   // NTTS[55] := 57;
   // NTTS[56] := 58;
   // NTTS[57] := 59;
   // NTTS[58] := 60;
   // NTTS[59] := 61;
   // NTTS[60] := 62;
   // NTTS[61] := 63;
   // NTTS[62] := 64;
   // NTTS[63] := 66;
   // SW_SQTS[2] := 1;
   // SW_SQTS[8] := 2;
   // SW_SQTS[9] := 2;
   // SW_SQTS[10] := 3;
   // SW_SQTS[11] := 3;
   // SW_SQTS[12] := 3;
   // SW_SQTS[13] := 3;
   // SW_SQTS[14] := 4;
   // SW_SQTS[15] := 4;
   // SW_SQTS[16] := 4;
   // SW_SQTS[17] := 4;
   // SW_SQTS[18] := 4;
   // SW_SQTS[19] := 4;
   // SW_SQTS[20] := 5;
   // SW_SQTS[21] := 5;
   // SW_SQTS[22] := 5;
   // SW_SQTS[23] := 2;
   // SW_SQTS[24] := 6;
   // SW_SQTS[25] := 6;
   // SW_SQTS[26] := 6;
   // SW_SQTS[27] := 6;
   // SW_SQTS[28] := 6;
   // SW_SQTS[29] := 6;
   // SW_SQTS[30] := 6;
   // SW_SQTS[31] := 6;
   // SWITCH[3] := 240;
   // SW_SQTS[36] := 7;
   // SW_SQTS[37] := 7;
   // SW_SQTS[38] := 7;
   // SW_SQTS[39] := 7;
   // SW_SQTS[40] := 7;
   // SW_SQTS[41] := 7;
   // SW_SQTS[42] := 7;
   // SW_SQTS[43] := 7;
   // SW_SQTS[44] := 7;
   // SW_SQTS[45] := 8;
   // SW_SQTS[46] := 8;
   // SW_SQTS[47] := 8;
   // SW_SQTS[48] := 8;
   // SW_SQTS[49] := 8;
   // SW_SQTS[50] := 8;
   // SW_SQTS[51] := 8;
   // SW_SQTS[52] := 8;
   // SW_SQTS[53] := 8;
   // SW_SQTS[54] := 8;
   // SW_SQTS[55] := 8;
   // SW_SQTS[56] := 8;
   // SW_SQTS[57] := 8;
   // SW_SQTS[58] := 8;
   // SW_SQTS[59] := 9;
   // SW_SQTS[60] := 9;
   // SW_SQTS[61] := 9;
   // SW_SQTS[62] := 9;
   // SW_SQTS[63] := 10;
   // SWITCH[0] := 252;
   // SWITCH[8] := 255;
   // SWITCH[4] := 167;
   // SWITCH[5] := 191;
   // SWITCH[6] := 252;
   // SWITCH[7] := 225;
   // SWITCH[2] := 255;
   // NSTT[48] := 47;
   // PTTS[27] := 34;
   // NSTT[38] := 37;
   // PTTS[30] := 31;
   // NTTS[1] := 3;
   // SWITCH[14] := 255;
   // ATAB[20] := 20;
   // PSTT[11] := 7;
   // NTTS[2] := 4;
   // PTTS[4] := 26;
   // PTTS[1] := 2;
   // NTTS[4] := 8;
   // SW_SQTS[1] := 1;
   // NSTT[26] := 4;
   // LSTT[48] := 255;
   // LSTT[63] := 255;
   // NSTT[63] := 62;
   // LSTT[61] := 255;
   // NSTT[61] := 60;
   // LSTT[64] := 1;
   // NSTT[64] := 1;
   // "Aux Reactor"."TIMER".MIX.PT := T#5M;
   // "Aux Reactor"."TIMER"."PRE-MIX".PT := T#5M;
   // SINI[6] := 255;
   // "Aux Reactor"."TIMER".TUBE.PT := T#5M;
   // "Aux Reactor"."TIMER".WASH.PT := T#5M;
   // SINI[5] := 255;
   // "Aux Reactor"."TIMER".REACTOR.PT := T#21.5H;
   // "Aux Reactor"."TIMER".PH_DELAY.PT := T#1M;
   // PTTS[29] := 30;
   // LSTT[37] := 255;
   // LSTT[25] := 24;
   // ATAB[19] := 19;
   // PSTT[15] := 11;
   // NSTT[37] := 36;
   // NSTT[25] := 24;
   // PTTS[28] := 28;
   // SW_SQTS[7] := 2;
   // SW_SQTS[6] := 2;
   // SW_SQTS[5] := 2;
   // SW_SQTS[4] := 2;
   // SWITCH[11] := 255;
   // SWITCH[13] := 239;
   // SWITCH[12] := 254;
   // PSTT[34] := 32;
   // PSTT[55] := 53;
   // PSTT[54] := 52;
   // LSTT[26] := 255;
   // SWITCH[10] := 239;
   // SWITCH[9] := 254;
   // SWITCH[1] := 231;
   // PTTS[2] := 3;
   // NSTT[49] := 48;
   // PSTT[53] := 51;
   // ATAB[0] := 1;
   // LSTT[49] := 255;
   // SINI[4] := 255;
   // SINI[2] := 255;
   // SW_SQTS[33] := 6;
   // SW_SQTS[32] := 6;
   // SINI[7] := 255;
   // SINI[8] := 255;
   // SINI[9] := 255;
   // LSTT[34] := 255;
   // LSTT[43] := 255;
   // PSTT[39] := 37;
   // NSTT[43] := 43;
   // LSTT[28] := 255;
   // LSTT[33] := 255;
   // ATAJ[66] := 66;
   // ATAB[66] := 66;
   // PSTT[66] := 63;
   // NSTT[33] := 26;
   // ASSJ[64] := 64;
   // ASSB[64] := 64;
   // PTTS[64] := 66;
   // NTTS[64] := 67;
   // SW_SQTS[64] := 10;
   // ATAJ[67] := 67;
   // ATAB[67] := 67;
   // PSTT[67] := 64;
   // NSTT[34] := 27;
   // LSTT[67] := 255;
   // ATAJ[68] := 68;
   // ATAB[68] := 68;
   // PSTT[68] := 65;
   // NSTT[67] := 65;
   // ASSJ[65] := 65;
   // ASSB[65] := 65;
   // PTTS[65] := 67;
   // NTTS[65] := 68;
   // SW_SQTS[65] := 10;
BEGIN
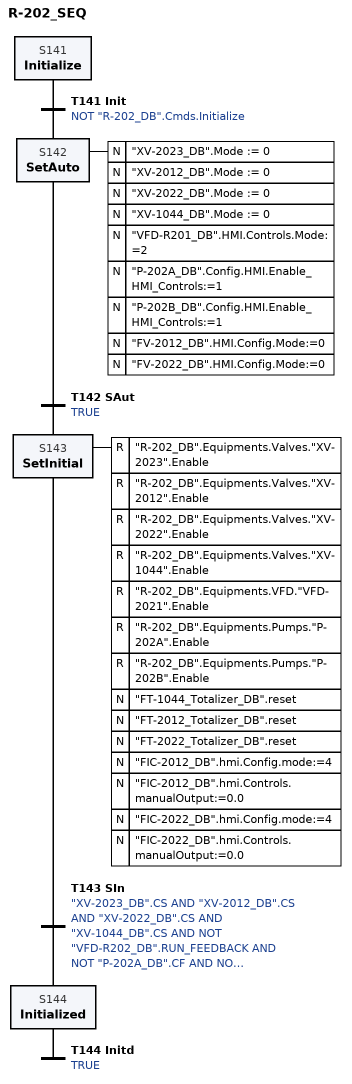
   // permanent pre-instructions
   NETWORK 1
      "R-202_Signals_FROM_T-101"();
      "R-202_Signals_FROM_T-102"();
      "R-202_Signals_FROM_T-103"();
      "R-202_Signals_FROM_T-104"();
      "R-202_SEQ_FC"();
      "R-202_Transitions_FC"();

   // sequencer 1
   STEP Initialize:   // S141, max time T#10S, warning time T#7S
   END_STEP
   TRANSITION Init FROM Initialize TO SetAuto   // T141
      := NOT "R-202_DB".Cmds.Initialize;
   END_TRANSITION
   STEP SetAuto:   // S142, max time T#10S, warning time T#7S
              N    "XV-2023_DB".Mode := 0
              N    "XV-2012_DB".Mode := 0
              N    "XV-2022_DB".Mode := 0
              N    "XV-1044_DB".Mode := 0
              N    "VFD-R201_DB".HMI.Controls.Mode:=2
              N    "P-202A_DB".Config.HMI.Enable_HMI_Controls:=1
              N    "P-202B_DB".Config.HMI.Enable_HMI_Controls:=1
              N    "FV-2012_DB".HMI.Config.Mode:=0
              N    "FV-2022_DB".HMI.Config.Mode:=0
   END_STEP
   TRANSITION SAut FROM SetAuto TO SetInitial   // T142
      := TRUE;
   END_TRANSITION
   STEP SetInitial:   // S143, max time T#10S, warning time T#7S
              R    "R-202_DB".Equipments.Valves."XV-2023".Enable
              R    "R-202_DB".Equipments.Valves."XV-2012".Enable
              R    "R-202_DB".Equipments.Valves."XV-2022".Enable
              R    "R-202_DB".Equipments.Valves."XV-1044".Enable
              R    "R-202_DB".Equipments.VFD."VFD-2021".Enable
              R    "R-202_DB".Equipments.Pumps."P-202A".Enable
              R    "R-202_DB".Equipments.Pumps."P-202B".Enable
              N    "FT-1044_Totalizer_DB".reset
              N    "FT-2012_Totalizer_DB".reset
              N    "FT-2022_Totalizer_DB".reset
              N    "FIC-2012_DB".hmi.Config.mode:=4
              N    "FIC-2012_DB".hmi.Controls.manualOutput:=0.0
              N    "FIC-2022_DB".hmi.Config.mode:=4
              N    "FIC-2022_DB".hmi.Controls.manualOutput:=0.0
   END_STEP
   TRANSITION SIn FROM SetInitial TO Initialized   // T143
      := "XV-2023_DB".CS AND "XV-2012_DB".CS AND "XV-2022_DB".CS AND "XV-1044_DB".CS AND NOT "VFD-R202_DB".RUN_FEEDBACK AND NOT "P-202A_DB".CF AND NOT "P-202B_DB".CF AND ("FV-2011_DB".CMD <= 0) AND ("FV-2021_DB".CMD <= 0) AND ("FT-1044_Totalizer_DB".Total = 0.0) AND ("FT-2012_Totalizer_DB".Total = 0.0) AND ("FT-2022_Totalizer_DB".Total = 0.0);
   END_TRANSITION
   STEP Initialized:   // S144, max time T#10S, warning time T#7S
      // Done Initialization
   END_STEP
   TRANSITION Initd FROM Initialized TO ?   // T144
      := TRUE;
   END_TRANSITION

   // permanent post-instructions
   NETWORK 1
      "R-202_FC_Outputs"();
END_FUNCTION_BLOCK

FUNCTION "R-202_FC_Outputs" : Void   // FC43, SCL
{ S7_Optimized_Access := 'TRUE' }
VERSION : 0.1
   VAR_TEMP
      Pump_A : Struct
         Cond_01 : Bool;   // Condition 01
         Cond_02 : Bool;
         Cond_03 : Bool;   // Condition 03
      END_STRUCT;
      Pump_B : Struct
         Cond_01 : Bool;   // Condition 01
         Cond_02 : Bool;   // Condition 02
         Cond_03 : Bool;   // Condition 03
      END_STRUCT;
      Motor : Struct
         Cond_01 : Bool;   // Condition 01
         Cond_02 : Bool;   // Condition 02
         Cond_03 : Bool;   // Condition 03
      END_STRUCT;
      XV : Struct
         "2023" : Bool;
         "2012" : Bool;
         "2022" : Bool;
         "1044" : Bool;
      END_STRUCT;
      "FV-2012" : Struct
         On : Bool;
         Cond_1 : Bool;
      END_STRUCT;
      "FV-2022" : Struct
         On : Bool;
         Cond_1 : Bool;
      END_STRUCT;
   END_VAR
BEGIN
   //****** Equipmens Activation*******
   //
   //**************************************************************
   //
   //IF "AlwaysFALSE" THEN
       //***********************************************Reactor Outlet Valve**********************************************************************
       IF "XV-2023_DB".Mode = 0 THEN
           "R-202_DB".Equipments.Valves."XV-2023".CmdOn := "R-202_DB".Equipments.Valves."XV-2023".Enable AND NOT "R-202_DB".Cmds.Hold;
           //Delay Off To avoid Overpressure the Lines
           #XV."2023" := "R-202_DB".Equipments.Valves."XV-2023".CmdOn;
           "R-202_Aux_DB".Timer."XV-2023".TOF(IN := #XV."2023",
                                              PT := "R-202_Aux_DB".Constants.CmdDelay);
           //Command to the Valve
           IF "R-202_Aux_DB".Timer."XV-2023".Q THEN
               "XV-2023_DB".CMD := 2;
           ELSE
               "XV-2023_DB".CMD := 1;
           END_IF;
           "R-202_DB".Equipments.Valves."XV-2023".TurningOff := NOT "R-202_DB".Equipments.Valves."XV-2023".CmdOn AND "R-202_Aux_DB".Timer."XV-2023".Q;
       END_IF;
       //***********************************************From T-101 Inlet Route********************************************************************
       IF "XV-2012_DB".Mode = 0 THEN
           "R-202_DB".Equipments.Valves."XV-2012".CmdOn := "R-202_DB".Equipments.Valves."XV-2012".Enable AND NOT "R-202_DB".Cmds.Hold;
           //Delay Off To avoid Overpressure the Lines
           #XV."2012" := "R-202_DB".Equipments.Valves."XV-2012".CmdOn;
           "R-202_Aux_DB".Timer."XV-2012".TOF(IN := #XV."2012",
                                              PT := "R-202_Aux_DB".Constants.CmdDelay);
           //Command to the Valve
           IF "R-202_Aux_DB".Timer."XV-2012".Q THEN
               "XV-2012_DB".CMD := 2;
           ELSE
               "XV-2012_DB".CMD := 1;
           END_IF;
           "R-202_DB".Equipments.Valves."XV-2012".TurningOff := NOT "R-202_DB".Equipments.Valves."XV-2012".CmdOn AND "R-202_Aux_DB".Timer."XV-2012".Q;
       END_IF;
       //***********************************************From T-102 Inlet Route********************************************************************
       IF "XV-2022_DB".Mode = 0 THEN
           "R-202_DB".Equipments.Valves."XV-2022".CmdOn := "R-202_DB".Equipments.Valves."XV-2022".Enable AND NOT "R-202_DB".Cmds.Hold;
           //Delay Off To avoid Overpressure the Lines
           #XV."2022" := "R-202_DB".Equipments.Valves."XV-2022".CmdOn;
           "R-202_Aux_DB".Timer."XV-2022".TOF(IN := #XV."2022",
                                              PT := "R-202_Aux_DB".Constants.CmdDelay);
           //Command to the Valve
           IF "R-202_Aux_DB".Timer."XV-2022".Q THEN
               "XV-2022_DB".CMD := 2;
           ELSE
               "XV-2022_DB".CMD := 1;
           END_IF;
           "R-202_DB".Equipments.Valves."XV-2022".TurningOff := NOT "R-202_DB".Equipments.Valves."XV-2022".CmdOn AND "R-202_Aux_DB".Timer."XV-2022".Q;
       END_IF;
       //***********************************************From T-104 Inlet Route (Water)********************************************************************
       IF "XV-1044_DB".Mode = 0 THEN
           "R-202_DB".Equipments.Valves."XV-1044".CmdOn := "R-202_DB".Equipments.Valves."XV-1044".Enable AND NOT "R-202_DB".Cmds.Hold;
           //Delay Off To avoid Overpressure the Lines
           #XV."1044" := "R-202_DB".Equipments.Valves."XV-1044".CmdOn;
           "R-202_Aux_DB".Timer."XV-1044".TOF(IN := #XV."1044",
                                              PT := "R-202_Aux_DB".Constants.CmdDelay);
           //Command to the Valve
           IF "R-202_Aux_DB".Timer."XV-1044".Q THEN
               "XV-1044_DB".CMD := 2;
           ELSE
               "XV-1044_DB".CMD := 1;
           END_IF;
           "R-202_DB".Equipments.Valves."XV-1044".TurningOff := NOT "R-202_DB".Equipments.Valves."XV-1044".CmdOn AND "R-202_Aux_DB".Timer."XV-2022".Q;
       END_IF;
       //***********************************************FIC-2012 Controller (From T-101)********************************************************************
       IF "FV-2012_DB".HMI.Config.Mode = 0 THEN
           #"FV-2012".Cond_1 := "R-202_DB".Equipments.Valves."FV-2012".Enable AND "XV-2012_DB".OS;
           "R-202_DB".Equipments.Valves."FV-2012".CmdOn := #"FV-2012".Cond_1 AND NOT "R-202_DB".Cmds.Hold AND NOT "R-202_DB".Status.Aborting;
           //Delay Off To avoid Overpressure the Lines
           #"FV-2012".On := "R-202_DB".Equipments.Valves."FV-2012".CmdOn;
           "R-202_Aux_DB".Timer."FV-2012".TOF(IN := #"FV-2012".On,
                                              PT := "R-202_Aux_DB".Constants.CmdDelay);
           IF "R-202_Aux_DB".Timer."FV-2012".Q THEN
               "FIC-2012_DB".enableManualMode := False;
               "FIC-2012_DB".enableRemoteSetpoint := False;
               "FIC-2012_DB".hmi.Controls.manualEnable := False;
               "FIC-2012_DB".hmi.Config.mode := 3;
           END_IF;     // ELSE
              // "FIC-2012_DB".enableManualMode := True;
              // "FIC-2012_DB".hmi.Controls.manualEnable := True;
              // "FIC-2012_DB".hmi.Config.mode := 4;
              // "FIC-2012_DB".hmi.Controls.manualOutput := 0;
         //  END_IF;
           "R-202_DB".Equipments.Valves."FV-2012".TurningOff := NOT "R-202_DB".Equipments.Valves."FV-2012".CmdOn AND "R-202_Aux_DB".Timer."FV-2012".Q;
       END_IF;
       //***********************************************FIC-2022 Controller (From T-102)********************************************************************
       IF "FV-2022_DB".HMI.Config.Mode = 0 THEN
           #"FV-2022".Cond_1 := "R-202_DB".Equipments.Valves."FV-2022".Enable AND "XV-2022_DB".OS;
           "R-202_DB".Equipments.Valves."FV-2022".CmdOn := #"FV-2022".Cond_1 AND NOT "R-202_DB".Cmds.Hold AND NOT "R-202_DB".Status.Aborting;
           //Delay Off To avoid Overpressure the Lines
           #"FV-2022".On := "R-202_DB".Equipments.Valves."FV-2022".CmdOn;
           "R-202_Aux_DB".Timer."FV-2022".TOF(IN := #"FV-2022".On,
                                              PT := "R-202_Aux_DB".Constants.CmdDelay);
           IF "R-202_Aux_DB".Timer."FV-2022".Q THEN

               IF "R-202_SEQ_DB".pH_Ctrl1.X OR "R-202_SEQ_DB".pH_Ctrl2.X OR "R-202_SEQ_DB".FillDone_T102.X THEN
                   //FIC-2022 Secondary Controller
                   "FIC-2022_DB".enableManualMode := False;
                   "FIC-2022_DB".hmi.Controls.manualEnable := False;
                   "FIC-2022_DB".enableRemoteSetpoint := true;
                   "FIC-2022_DB".hmi.Config.mode := 6;

                   //PHIC-R-202 pH Primary Controller
                   "PHIC-R-202_DB".enableRemoteSetpoint := False;
                   "PHIC-R-202_DB".enableManualMode := False;
                   "PHIC-R-202_DB".hmi.Controls.manualEnable := False;
                   "PHIC-R-202_DB".hmi.Config.mode := 3;
               ELSIF "R-202_SEQ_DB".Y.X THEN
                   //FIC-2022 Secondary Controller
                   "FIC-2022_DB".enableManualMode := False;
                   "FIC-2022_DB".hmi.Controls.manualEnable := False;
                   "FIC-2022_DB".enableRemoteSetpoint := false;
                   "FIC-2022_DB".hmi.Config.mode := 3;

                   //PHIC-R-202 pH Primary Controller
                   "PHIC-R-202_DB".enableRemoteSetpoint := False;
                   "PHIC-R-202_DB".enableManualMode := False;
                   "PHIC-R-202_DB".hmi.Controls.manualEnable := False;
                   "PHIC-R-202_DB".hmi.Config.mode := 3;

               END_IF;



           END_IF;     // ELSE
               //FIC-2022 Secondary Controller
             //  "FIC-2022_DB".enableManualMode := True;
             //  "FIC-2022_DB".hmi.Controls.manualEnable := True;
             //  "FIC-2022_DB".enableRemoteSetpoint := False;
             //  "FIC-2022_DB".hmi.Config.mode := 4;
             //  "FIC-2022_DB".hmi.Controls.manualOutput := 0;

               //PHIC-R-202 pH Primary  Controller
             //  "PHIC-R-202_DB".enableManualMode := True;
             //  "PHIC-R-202_DB".hmi.Controls.manualEnable := True;
             //  "PHIC-R-202_DB".enableRemoteSetpoint := False;
             //  "PHIC-R-202_DB".hmi.Config.mode := 4;
            //   "PHIC-R-202_DB".hmi.Controls.manualOutput := 0;
         //  END_IF;
           "R-202_DB".Equipments.Valves."FV-2022".TurningOff := NOT "R-202_DB".Equipments.Valves."FV-2022".CmdOn AND "R-202_Aux_DB".Timer."FV-2022".Q;
       END_IF;
       //***********************************************Recirculate/Feed Pump A********************************************************************
       // Condition to CmdOn "On Command" 
       IF "P-202A_DB".Config.HMI.Enable_HMI_Controls = 1 THEN
           #Pump_A.Cond_01 := "R-202_DB".Equipments.Pumps."P-202A".Enable AND ("R-202_DB".PmpSel."P-202AB" = 1 OR "R-202_DB".PmpSel."P-202AB" = 3);
           #Pump_A.Cond_02 := "XV-2023_DB".OS AND "R-202_Read_FROM_T-103_DB".RouteOpened; //Route Open to sent to the T-103 (Cooling Tank)
           "R-202_DB".Equipments.Pumps."P-202A".CmdOn := #Pump_A.Cond_01 AND #Pump_A.Cond_02 AND NOT "R-202_DB".Cmds.Hold;
           IF "R-202_DB".Equipments.Pumps."P-202A".CmdOn THEN
               "P-202A_DB".Stop_CMD := False;
               "P-202A_DB".Start_CMD := true;
               "P-202A_DB".ON := TRUE;
               "P-202A_DB".OFF := FALSE;
           ELSE
               "P-202A_DB".Stop_CMD := TRUE;
               "P-202A_DB".Start_CMD := FALSE;
               "P-202A_DB".ON := FALSE;
               "P-202A_DB".OFF := TRUE;
           END_IF;
       END_IF;
       //***********************************************Recirculate/Feed Pump B********************************************************************
       // Condition to CmdOn "On Command" 
       IF "P-202B_DB".Config.HMI.Enable_HMI_Controls = 1 THEN
           #Pump_B.Cond_01 := "R-202_DB".Equipments.Pumps."P-202B".Enable AND ("R-202_DB".PmpSel."P-202AB" = 2 OR "R-202_DB".PmpSel."P-202AB" = 3);
           #Pump_B.Cond_02 := "XV-2023_DB".OS AND "R-202_Read_FROM_T-103_DB".RouteOpened; //Route Open to sent to the T-103 (Cooling Tank)
           "R-202_DB".Equipments.Pumps."P-202B".CmdOn := #Pump_B.Cond_01 AND #Pump_B.Cond_02  AND NOT "R-202_DB".Cmds.Hold;
           IF "R-202_DB".Equipments.Pumps."P-202B".CmdOn THEN
               "P-202B_DB".Stop_CMD := False;
               "P-202B_DB".Start_CMD := true;
               "P-202B_DB".ON := TRUE;
               "P-202B_DB".OFF := FALSE;
           ELSE
               "P-202B_DB".Stop_CMD := TRUE;
               "P-202B_DB".Start_CMD := FALSE;
               "P-202B_DB".ON := FALSE;
               "P-202B_DB".OFF := TRUE;
           END_IF;
       END_IF;
       //***********************************************Mixer********************************************************************
       IF "VFD-R202_DB".HMI.Controls.Mode = 2 THEN
           "R-202_Aux_DB"."Real"."VFD-R202".Start := (("LT-2021_DB".SAI > "R-202_Recipe".MinLevelMixerOn + 2.0) OR "R-202_Aux_DB"."Real"."VFD-R202".Start) AND NOT "R-202_Aux_DB"."Real"."VFD-R202".Stop;
           "R-202_Aux_DB"."Real"."VFD-R202".Stop := ("LT-2021_DB".SAI < "R-202_Recipe".MinLevelMixerOn - 1.0);
           #Motor.Cond_01 := "R-202_DB".Equipments.VFD."VFD-2021".Enable AND "LT-2021_DB".SAI > "R-202_Recipe".MinLevelMixerOn;
           "R-202_DB".Equipments.VFD."VFD-2021".CmdOn := #Motor.Cond_01 AND NOT "R-202_DB".Cmds.Hold AND NOT "R-202_DB".Status.Aborting;;
           IF "R-202_DB".Equipments.VFD."VFD-2021".CmdOn THEN
               "VFD-R202_DB".PLCCommand := TRUE;
           ELSE
               "VFD-R202_DB".PLCCommand := FALSE;
           END_IF;
       END_IF;
   //END_IF;

   //***************Interlocks to T-103***************//
   //Transfering
   "R-202_Write_TO_T-103_DB".Transfering := ("XV-2023_DB".OS) AND (("P-202A_DB".CF AND ("PT-202A_DB".SAI > 0.2)) OR ("P-202B_DB".CF AND ("PT-202B_DB".SAI > 0.2)));
   "R-202_Write_TO_T-103_DB"."Transfer_To_T-103_Done" := "R-202_DB".Status.Step = 66;// AND "XV-2023_DB".CS AND NOT "P-202A_DB".CF AND NOT "P-202B_DB".CF AND NOT "VFD-R202_DB".RUN_FEEDBACK;
   //***************Interlocks to T-101***************//
   "R-202_Write_TO_T-101_DB".OpenRoute := "XV-2012_DB".OS AND ("FV-2012_DB".CMD > 0);
   "R-202_Write_TO_T-101_DB".RouteOpened := "XV-2012_DB".OS AND ("FV-2012_DB".CMD > 0);

   //***************Interlocks to T-102***************//
   "R-202_Write_TO_T-102_DB".OpenRoute := "XV-2022_DB".OS AND ("FV-2022_DB".CMD > 0);
   "R-202_Write_TO_T-102_DB".RouteOpened := "XV-2022_DB".OS AND ("FV-2022_DB".CMD > 0);
   //***************Abort Signals***************//
   //******Abort T-101*****//
   IF "R-202_DB".Status.Aborting THEN

       "R-202_Write_TO_T-101_DB".Abort := "R-202_SEQ_DB".S_NO >= 21 AND "R-202_SEQ_DB".S_NO <= 39;
       "R-202_Write_TO_T-102_DB".Abort := "R-202_SEQ_DB".S_NO >= 21 AND "R-202_SEQ_DB".S_NO <= 39;
       "R-202_Write_TO_T-103_DB".Abort :=("R-202_DB".Status.State = 3);

   END_IF;

   //***************Interlocks to T-104***************//
   "R-202_Write_TO_T-104_DB".ReqWater := "XV-2023_DB".CS AND "XV-1044_DB".OS AND ("R-202_DB".Status.Step = 23 OR "R-202_DB".Status.Step = 68 OR "R-202_DB".Status.Step = 66);

   //***************Valves Status***************//
   "R-202_Aux_DB"."Bool".TOff := "R-202_DB".Equipments.Valves."XV-2023".TurningOff OR "R-202_DB".Equipments.Valves."XV-2012".TurningOff OR "R-202_DB".Equipments.Valves."XV-2022".TurningOff OR "R-202_DB".Equipments.Valves."XV-1044".TurningOff;
   //***************Timers***************//
   //Pre-Mix Timer
   "R-202_Aux_DB"."Bool".PreMixT_En := "R-202_DB".Status.Step = 26 AND "R-202_Read_FROM_T-102_DB".Recirculating AND "R-202_Read_FROM_T-101_DB".Recirculating; //T-102 AND T-102 Mixing
   "R-202_Aux_DB"."Bool".PreMixT_Reset := "R-202_DB".Cmds.Abort OR "R-202_DB".Status.Step = 1;
   //pH Stabilize Timer
   "R-202_Aux_DB"."Bool".StabpHTEn := "R-202_Aux_DB"."Bool".StabpHTEnStep AND "FT-2022_DB".SAI > 0.2 AND "FT-2012_DB".SAI > 0.2;
   "R-202_Aux_DB"."Bool".StabpHTEn_Reset := "R-202_DB".Cmds.Abort OR "R-202_DB".Status.Step = 1;
   //Reaction Timer
   "R-202_Aux_DB"."Bool".ReactorTEn := "R-202_DB".Status.Step = 40;
   "R-202_Aux_DB"."Bool".ReactorT_Reset := "R-202_DB".Cmds.Abort OR "R-202_DB".Status.Step = 1;
   //Last Run Timer
   "R-202_Aux_DB"."Bool".FlushOutTEn := ("R-202_DB".Status.Step = 67 OR "R-202_DB".Status.Step = 64) AND ("P-202A_DB".CF OR "P-202B_DB".CF) AND "XV-2023_DB".OS;
   //Mix To Clean Timer
   "R-202_Aux_DB"."Bool".MixToCleanTEn := "R-202_DB".Status.Step = 63 AND "VFD-R202_DB".RUN_FEEDBACK;
   "R-202_Aux_DB"."Bool".MixToCleanT_Reset := "R-202_DB".Cmds.Abort OR "R-202_DB".Status.Step = 1;
END_FUNCTION

FUNCTION "R-202_SEQ_FC" : Void   // FC77, LAD
{ S7_Optimized_Access := 'TRUE' }
VERSION : 0.1
   VAR_TEMP   // added for the SCL form of the ladder/FBD networks
      _w1 : Bool;
      _w2 : Bool;
   END_VAR
BEGIN

REGION Network 2: Abort
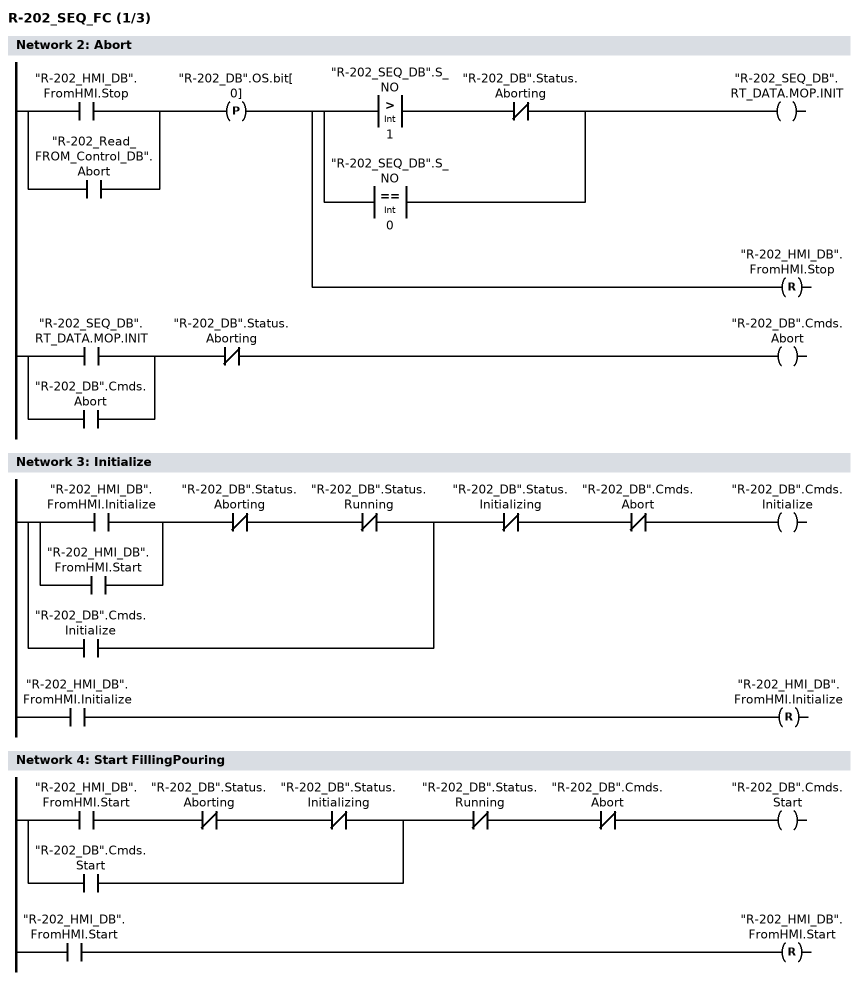
   RUNG wire#powerrail
      Contact( "R-202_HMI_DB".FromHMI.Stop )
      wire#w1
      P_Trig( "R-202_DB".OS.bit[0] )
      wire#w2
      { S7_Templates := "SrcType := Int" } GT_Contact(in1 := "R-202_SEQ_DB".S_NO, in2 := 1)
      I_Contact( "R-202_DB".Status.Aborting )
      wire#w3
      Coil( "R-202_SEQ_DB".RT_DATA.MOP.INIT )
   END_RUNG
   RUNG wire#powerrail
      Contact( "R-202_Read_FROM_Control_DB".Abort )
   END_RUNG wire#w1
   RUNG wire#w2
      { S7_Templates := "SrcType := Int" } EQ_Contact(in1 := "R-202_SEQ_DB".S_NO, in2 := 0)
   END_RUNG wire#w3
   RUNG wire#w2
      R_Coil( "R-202_HMI_DB".FromHMI.Stop )
   END_RUNG
   RUNG wire#powerrail
      Contact( "R-202_SEQ_DB".RT_DATA.MOP.INIT )
      wire#w4
      I_Contact( "R-202_DB".Status.Aborting )
      Coil( "R-202_DB".Cmds.Abort )
   END_RUNG
   RUNG wire#powerrail
      Contact( "R-202_DB".Cmds.Abort )
   END_RUNG wire#w4
   // the same network as SCL:
   #_w1 := "R-202_HMI_DB".FromHMI.Stop OR "R-202_Read_FROM_Control_DB".Abort;
   #_w2 := #_w1 AND NOT "R-202_DB".OS.bit[0];   // rising edge
   "R-202_DB".OS.bit[0] := #_w1;
   "R-202_SEQ_DB".RT_DATA.MOP.INIT := #_w2 AND ((("R-202_SEQ_DB".S_NO > 1) AND NOT "R-202_DB".Status.Aborting) OR ("R-202_SEQ_DB".S_NO = 0));
   IF #_w2 THEN "R-202_HMI_DB".FromHMI.Stop := FALSE; END_IF;
   "R-202_DB".Cmds.Abort := ("R-202_SEQ_DB".RT_DATA.MOP.INIT OR "R-202_DB".Cmds.Abort) AND NOT "R-202_DB".Status.Aborting;
END_REGION

REGION Network 3: Initialize
   RUNG wire#powerrail
      Contact( "R-202_HMI_DB".FromHMI.Initialize )
      wire#w1
      I_Contact( "R-202_DB".Status.Aborting )
      I_Contact( "R-202_DB".Status.Running )
      wire#w2
      I_Contact( "R-202_DB".Status.Initializing )
      I_Contact( "R-202_DB".Cmds.Abort )
      Coil( "R-202_DB".Cmds.Initialize )
   END_RUNG
   RUNG wire#powerrail
      Contact( "R-202_HMI_DB".FromHMI.Start )
   END_RUNG wire#w1
   RUNG wire#powerrail
      Contact( "R-202_DB".Cmds.Initialize )
   END_RUNG wire#w2
   RUNG wire#powerrail
      Contact( "R-202_HMI_DB".FromHMI.Initialize )
      R_Coil( "R-202_HMI_DB".FromHMI.Initialize )
   END_RUNG
   // the same network as SCL:
   "R-202_DB".Cmds.Initialize := ((("R-202_HMI_DB".FromHMI.Initialize OR "R-202_HMI_DB".FromHMI.Start) AND NOT "R-202_DB".Status.Aborting AND NOT "R-202_DB".Status.Running) OR "R-202_DB".Cmds.Initialize) AND NOT "R-202_DB".Status.Initializing AND NOT "R-202_DB".Cmds.Abort;
   IF "R-202_HMI_DB".FromHMI.Initialize THEN "R-202_HMI_DB".FromHMI.Initialize := FALSE; END_IF;
END_REGION

REGION Network 4: Start FillingPouring
   RUNG wire#powerrail
      Contact( "R-202_HMI_DB".FromHMI.Start )
      I_Contact( "R-202_DB".Status.Aborting )
      I_Contact( "R-202_DB".Status.Initializing )
      wire#w1
      I_Contact( "R-202_DB".Status.Running )
      I_Contact( "R-202_DB".Cmds.Abort )
      Coil( "R-202_DB".Cmds.Start )
   END_RUNG
   RUNG wire#powerrail
      Contact( "R-202_DB".Cmds.Start )
   END_RUNG wire#w1
   RUNG wire#powerrail
      Contact( "R-202_HMI_DB".FromHMI.Start )
      R_Coil( "R-202_HMI_DB".FromHMI.Start )
   END_RUNG
   // the same network as SCL:
   "R-202_DB".Cmds.Start := (("R-202_HMI_DB".FromHMI.Start AND NOT "R-202_DB".Status.Aborting AND NOT "R-202_DB".Status.Initializing) OR "R-202_DB".Cmds.Start) AND NOT "R-202_DB".Status.Running AND NOT "R-202_DB".Cmds.Abort;
   IF "R-202_HMI_DB".FromHMI.Start THEN "R-202_HMI_DB".FromHMI.Start := FALSE; END_IF;
END_REGION

REGION Network 5: Procedure Selected
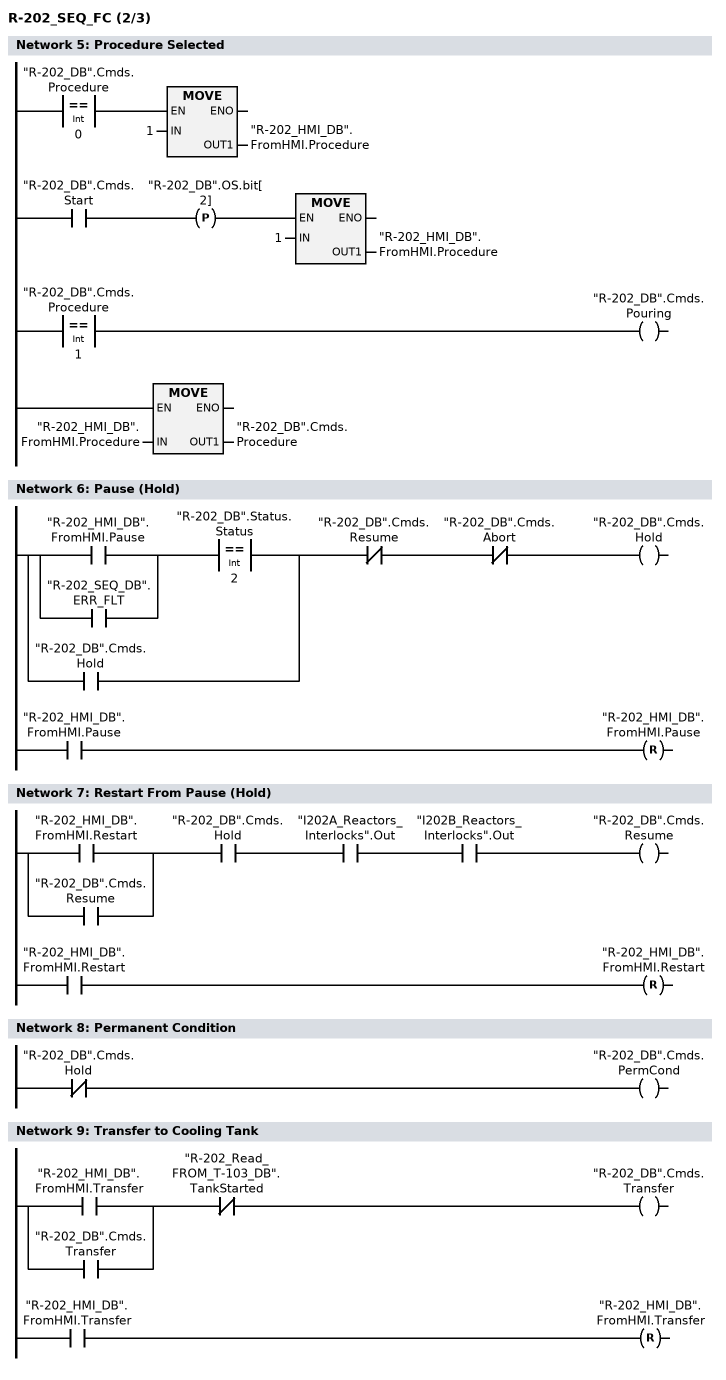
   RUNG wire#powerrail
      { S7_Templates := "SrcType := Int" } EQ_Contact(in1 := "R-202_DB".Cmds.Procedure, in2 := 0)
      Move(in := 1, out1 => "R-202_HMI_DB".FromHMI.Procedure)
   END_RUNG
   RUNG wire#powerrail
      Contact( "R-202_DB".Cmds.Start )
      P_Trig( "R-202_DB".OS.bit[2] )
      Move(in := 1, out1 => "R-202_HMI_DB".FromHMI.Procedure)
   END_RUNG
   RUNG wire#powerrail
      { S7_Templates := "SrcType := Int" } EQ_Contact(in1 := "R-202_DB".Cmds.Procedure, in2 := 1)
      Coil( "R-202_DB".Cmds.Pouring )
   END_RUNG
   RUNG wire#powerrail
      Move(in := "R-202_HMI_DB".FromHMI.Procedure, out1 => "R-202_DB".Cmds.Procedure)
   END_RUNG
   // the same network as SCL:
   IF "R-202_DB".Cmds.Procedure = 0 THEN "R-202_HMI_DB".FromHMI.Procedure := 1; END_IF;
   #_w1 := "R-202_DB".Cmds.Start AND NOT "R-202_DB".OS.bit[2];   // rising edge
   "R-202_DB".OS.bit[2] := "R-202_DB".Cmds.Start;
   IF #_w1 THEN "R-202_HMI_DB".FromHMI.Procedure := 1; END_IF;
   "R-202_DB".Cmds.Pouring := "R-202_DB".Cmds.Procedure = 1;
   "R-202_DB".Cmds.Procedure := "R-202_HMI_DB".FromHMI.Procedure;
END_REGION

REGION Network 6: Pause (Hold)
   RUNG wire#powerrail
      Contact( "R-202_HMI_DB".FromHMI.Pause )
      wire#w1
      { S7_Templates := "SrcType := Int" } EQ_Contact(in1 := "R-202_DB".Status.Status, in2 := 2)
      wire#w2
      I_Contact( "R-202_DB".Cmds.Resume )
      I_Contact( "R-202_DB".Cmds.Abort )
      Coil( "R-202_DB".Cmds.Hold )
   END_RUNG
   RUNG wire#powerrail
      Contact( "R-202_SEQ_DB".ERR_FLT )
   END_RUNG wire#w1
   RUNG wire#powerrail
      Contact( "R-202_DB".Cmds.Hold )
   END_RUNG wire#w2
   RUNG wire#powerrail
      Contact( "R-202_HMI_DB".FromHMI.Pause )
      R_Coil( "R-202_HMI_DB".FromHMI.Pause )
   END_RUNG
   // the same network as SCL:
   "R-202_DB".Cmds.Hold := ((("R-202_HMI_DB".FromHMI.Pause OR "R-202_SEQ_DB".ERR_FLT) AND ("R-202_DB".Status.Status = 2)) OR "R-202_DB".Cmds.Hold) AND NOT "R-202_DB".Cmds.Resume AND NOT "R-202_DB".Cmds.Abort;
   IF "R-202_HMI_DB".FromHMI.Pause THEN "R-202_HMI_DB".FromHMI.Pause := FALSE; END_IF;
END_REGION

REGION Network 7: Restart From Pause (Hold)
   RUNG wire#powerrail
      Contact( "R-202_HMI_DB".FromHMI.Restart )
      wire#w1
      Contact( "R-202_DB".Cmds.Hold )
      Contact( "I202A_Reactors_Interlocks".Out )
      Contact( "I202B_Reactors_Interlocks".Out )
      Coil( "R-202_DB".Cmds.Resume )
   END_RUNG
   RUNG wire#powerrail
      Contact( "R-202_DB".Cmds.Resume )
   END_RUNG wire#w1
   RUNG wire#powerrail
      Contact( "R-202_HMI_DB".FromHMI.Restart )
      R_Coil( "R-202_HMI_DB".FromHMI.Restart )
   END_RUNG
   // the same network as SCL:
   "R-202_DB".Cmds.Resume := ("R-202_HMI_DB".FromHMI.Restart OR "R-202_DB".Cmds.Resume) AND "R-202_DB".Cmds.Hold AND "I202A_Reactors_Interlocks".Out AND "I202B_Reactors_Interlocks".Out;
   IF "R-202_HMI_DB".FromHMI.Restart THEN "R-202_HMI_DB".FromHMI.Restart := FALSE; END_IF;
END_REGION

REGION Network 8: Permanent Condition
   RUNG wire#powerrail
      I_Contact( "R-202_DB".Cmds.Hold )
      Coil( "R-202_DB".Cmds.PermCond )
   END_RUNG
   // the same network as SCL:
   "R-202_DB".Cmds.PermCond := NOT "R-202_DB".Cmds.Hold;
END_REGION

REGION Network 9: Transfer to Cooling Tank
   RUNG wire#powerrail
      Contact( "R-202_HMI_DB".FromHMI.Transfer )
      wire#w1
      I_Contact( "R-202_Read_FROM_T-103_DB".TankStarted )
      Coil( "R-202_DB".Cmds.Transfer )
   END_RUNG
   RUNG wire#powerrail
      Contact( "R-202_DB".Cmds.Transfer )
   END_RUNG wire#w1
   RUNG wire#powerrail
      Contact( "R-202_HMI_DB".FromHMI.Transfer )
      R_Coil( "R-202_HMI_DB".FromHMI.Transfer )
   END_RUNG
   // the same network as SCL:
   "R-202_DB".Cmds.Transfer := ("R-202_HMI_DB".FromHMI.Transfer OR "R-202_DB".Cmds.Transfer) AND NOT "R-202_Read_FROM_T-103_DB".TankStarted;
   IF "R-202_HMI_DB".FromHMI.Transfer THEN "R-202_HMI_DB".FromHMI.Transfer := FALSE; END_IF;
END_REGION

REGION Network 10: Tank Wash
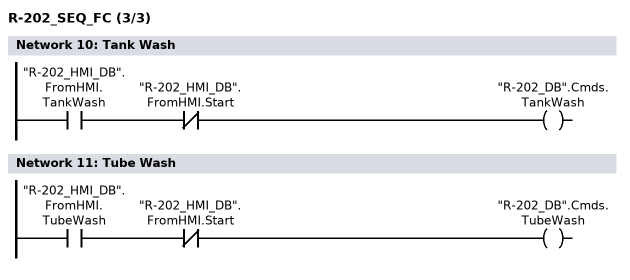
   RUNG wire#powerrail
      Contact( "R-202_HMI_DB".FromHMI.TankWash )
      I_Contact( "R-202_HMI_DB".FromHMI.Start )
      Coil( "R-202_DB".Cmds.TankWash )
   END_RUNG
   // the same network as SCL:
   "R-202_DB".Cmds.TankWash := "R-202_HMI_DB".FromHMI.TankWash AND NOT "R-202_HMI_DB".FromHMI.Start;
END_REGION

REGION Network 11: Tube Wash
   RUNG wire#powerrail
      Contact( "R-202_HMI_DB".FromHMI.TubeWash )
      I_Contact( "R-202_HMI_DB".FromHMI.Start )
      Coil( "R-202_DB".Cmds.TubeWash )
   END_RUNG
   // the same network as SCL:
   "R-202_DB".Cmds.TubeWash := "R-202_HMI_DB".FromHMI.TubeWash AND NOT "R-202_HMI_DB".FromHMI.Start;
END_REGION

REGION Network 12 (SCL): Sequence Status
   IF "R-202_SEQ_DB".S_NO = 1 THEN
       "R-202_DB".Status.Status := 1; //Idle
   ELSIF ("R-202_SEQ_DB".S_NO > 1 AND "R-202_SEQ_DB".S_NO <= 150)  AND NOT "R-202_SEQ_DB".ERR_FLT AND NOT "R-202_DB".Cmds.Hold THEN
       "R-202_DB".Status.Status := 2; //Running
   ELSIF "R-202_SEQ_DB".S_NO >= 151 AND "R-202_SEQ_DB".S_NO <= 160 AND NOT "R-202_SEQ_DB".ERR_FLT THEN
       "R-202_DB".Status.Status := 3; // Stopping
   ELSIF "R-202_SEQ_DB".ERR_FLT  AND ("R-202_SEQ_DB".S_NO > 1 AND "R-202_SEQ_DB".S_NO <= 150) THEN
       "R-202_DB".Status.Status := 4; //Held
   ELSIF  "R-202_SEQ_DB".ERR_FLT AND  ("R-202_SEQ_DB".S_NO > 1 AND "R-202_SEQ_DB".S_NO <= 150) AND "R-202_Aux_DB"."Bool".TOff  THEN
       "R-202_DB".Status.Status := 5; // Holding
   ELSE
       "R-202_DB".Status.Status := 6; // Unknown
   END_IF;

   "R-202_DB".Status.Running := ("R-202_SEQ_DB".S_NO > 3 AND "R-202_SEQ_DB".S_NO <= 150);
   "R-202_DB".Status.Initializing := ("R-202_SEQ_DB".S_NO >= 141 AND "R-202_SEQ_DB".S_NO <= 150);
   //Enable/Disable HMI Start/Stop Button
   "R-202_HMI_DB".ToHMI.EnStopButton:=("R-202_DB".Status.Status>1) OR "R-202_DB".Status.Step=0; //Enable HMI Stop Button
   "R-202_HMI_DB".ToHMI.EnStartButton := "R-202_DB".Status.Status = 1;     //Enable Start Button
   "R-202_HMI_DB".ToHMI.EnPauseButton := "R-202_DB".Status.Status = 2 ; //Enable Pause Button
   "R-202_HMI_DB".ToHMI.EnRestartButton := "R-202_DB".Status.Status = 4; //Enable Restart Button

   //****Interlock Activated
   "R-202_HMI_DB".ToHMI.InterlockActivated := "I202A_Reactors_Interlocks".Out AND "I202B_Reactors_Interlocks".Out;
END_REGION

REGION Network 13 (SCL): Sequence Step
   "R-202_DB".Status.Step := "R-202_SEQ_DB".S_NO;
END_REGION

REGION Network 14 (SCL): Sequence state (Procedure running)
   IF "R-202_SEQ_DB".S_NO = 3 OR "R-202_SEQ_DB".S_NO = 4 THEN
       "R-202_DB".Status.State := 1; //Seq Selection
   ELSIF "R-202_SEQ_DB".S_NO >= 21 AND "R-202_SEQ_DB".S_NO <= 60 THEN
       "R-202_DB".Status.State := 2; //Pouring 
   ELSIF "R-202_SEQ_DB".S_NO >= 61 AND "R-202_SEQ_DB".S_NO <= 80 THEN
       "R-202_DB".Status.State := 3; //Transfering
   ELSIF "R-202_SEQ_DB".S_NO >= 81 AND "R-202_SEQ_DB".S_NO <= 100 THEN
       "R-202_DB".Status.State := 4; //Washing Tank
   ELSIF "R-202_SEQ_DB".S_NO >= 101 AND "R-202_SEQ_DB".S_NO <= 140 THEN
       "R-202_DB".Status.State := 5; //Washing Lines
   ELSIF "R-202_SEQ_DB".S_NO >= 151 AND "R-202_SEQ_DB".S_NO <= 160 THEN
       "R-202_DB".Status.State := 6; //Aborting
   ELSIF "R-202_SEQ_DB".S_NO >= 141 AND "R-202_SEQ_DB".S_NO <= 150 THEN
       "R-202_DB".Status.State := 7; //Initializing
   ELSE
       "R-202_DB".Status.State := 0;
   END_IF;
END_REGION
END_FUNCTION

FUNCTION "R-202_Transitions_FC" : Void   // FC80, SCL
{ S7_Optimized_Access := 'TRUE' }
VERSION : 0.1
BEGIN

   //*****"Transition" for Low Level and Low pressure meaning "Tank is Empty"
   "R-202_Aux_DB"."Bool".Transitions.TankEmpty := "LT-2021_DB".SAI <= "ReactorLowLevelSetpoint" AND (("PT-202A_DB".SAI <= 1.0) AND ("PT-202B_DB".SAI <= 1.0));
END_FUNCTION

